                      InputLimitSwitchClosed := "20_TANKS_IP_DATA".RIO_05.SECOND_TANK.TANK_VENT_A_CLSD,
                      Open => "1092_HMI_OP_FLAGS".CV427_428_PVVA_Alarms[11].Open,
                      Closed => "1092_HMI_OP_FLAGS".CV427_428_PVVA_Alarms[11].Closed,
                      Moving => "1092_HMI_OP_FLAGS".CV427_428_PVVA_Alarms[11].Moving,
                      Fault => "1092_HMI_OP_FLAGS".CV427_428_PVVA_Alarms[11].Fault);
END_REGION

REGION Network 6: 600-CV-427, 600-CV-428 Alarms (RIO 06: 6P, 6S)
   RUNG wire#powerrail
      "1603_VALVE_STATE"(InputLimitSwitchOpen := "20_TANKS_IP_DATA".RIO_06.FIRST_TANK.TANK_VENT_A_OPEN, InputLimitSwitchClosed := "20_TANKS_IP_DATA".RIO_06.FIRST_TANK.TANK_VENT_A_CLSD, Open => "1092_HMI_OP_FLAGS".CV427_428_PVVA_Alarms[12].Open, Closed => "1092_HMI_OP_FLAGS".CV427_428_PVVA_Alarms[12].Closed, Moving => "1092_HMI_OP_FLAGS".CV427_428_PVVA_Alarms[12].Moving, Fault => "1092_HMI_OP_FLAGS".CV427_428_PVVA_Alarms[12].Fault)
   END_RUNG
   RUNG wire#powerrail
      "1603_VALVE_STATE"(InputLimitSwitchOpen := "20_TANKS_IP_DATA".RIO_06.SECOND_TANK.TANK_VENT_A_OPEN, InputLimitSwitchClosed := "20_TANKS_IP_DATA".RIO_06.SECOND_TANK.TANK_VENT_A_CLSD, Open => "1092_HMI_OP_FLAGS".CV427_428_PVVA_Alarms[13].Open, Closed => "1092_HMI_OP_FLAGS".CV427_428_PVVA_Alarms[13].Closed, Moving => "1092_HMI_OP_FLAGS".CV427_428_PVVA_Alarms[13].Moving, Fault => "1092_HMI_OP_FLAGS".CV427_428_PVVA_Alarms[13].Fault)
   END_RUNG
   // the same network as SCL:
   "1603_VALVE_STATE"(InputLimitSwitchOpen := "20_TANKS_IP_DATA".RIO_06.FIRST_TANK.TANK_VENT_A_OPEN,
                      InputLimitSwitchClosed := "20_TANKS_IP_DATA".RIO_06.FIRST_TANK.TANK_VENT_A_CLSD,
                      Open => "1092_HMI_OP_FLAGS".CV427_428_PVVA_Alarms[12].Open,
                      Closed => "1092_HMI_OP_FLAGS".CV427_428_PVVA_Alarms[12].Closed,
                      Moving => "1092_HMI_OP_FLAGS".CV427_428_PVVA_Alarms[12].Moving,
                      Fault => "1092_HMI_OP_FLAGS".CV427_428_PVVA_Alarms[12].Fault);
   "1603_VALVE_STATE"(InputLimitSwitchOpen := "20_TANKS_IP_DATA".RIO_06.SECOND_TANK.TANK_VENT_A_OPEN,
                      InputLimitSwitchClosed := "20_TANKS_IP_DATA".RIO_06.SECOND_TANK.TANK_VENT_A_CLSD,
                      Open => "1092_HMI_OP_FLAGS".CV427_428_PVVA_Alarms[13].Open,
                      Closed => "1092_HMI_OP_FLAGS".CV427_428_PVVA_Alarms[13].Closed,
                      Moving => "1092_HMI_OP_FLAGS".CV427_428_PVVA_Alarms[13].Moving,
                      Fault => "1092_HMI_OP_FLAGS".CV427_428_PVVA_Alarms[13].Fault);
END_REGION

REGION Network 7: 600-CV-427, 600-CV-428 Alarms (RIO 07: APT)
   RUNG wire#powerrail
      "1603_VALVE_STATE"(InputLimitSwitchOpen := "20_TANKS_IP_DATA".RIO_07.FIRST_TANK.TANK_VENT_A_OPEN, InputLimitSwitchClosed := "20_TANKS_IP_DATA".RIO_07.FIRST_TANK.TANK_VENT_A_CLSD, Open => "1092_HMI_OP_FLAGS".CV427_428_PVVA_Alarms[14].Open, Closed => "1092_HMI_OP_FLAGS".CV427_428_PVVA_Alarms[14].Closed, Moving => "1092_HMI_OP_FLAGS".CV427_428_PVVA_Alarms[14].Moving, Fault => "1092_HMI_OP_FLAGS".CV427_428_PVVA_Alarms[14].Fault)
   END_RUNG
   // the same network as SCL:
   "1603_VALVE_STATE"(InputLimitSwitchOpen := "20_TANKS_IP_DATA".RIO_07.FIRST_TANK.TANK_VENT_A_OPEN,
                      InputLimitSwitchClosed := "20_TANKS_IP_DATA".RIO_07.FIRST_TANK.TANK_VENT_A_CLSD,
                      Open => "1092_HMI_OP_FLAGS".CV427_428_PVVA_Alarms[14].Open,
                      Closed => "1092_HMI_OP_FLAGS".CV427_428_PVVA_Alarms[14].Closed,
                      Moving => "1092_HMI_OP_FLAGS".CV427_428_PVVA_Alarms[14].Moving,
                      Fault => "1092_HMI_OP_FLAGS".CV427_428_PVVA_Alarms[14].Fault);
END_REGION
END_FUNCTION

FUNCTION "1087_600CV429_430_STATUS" : Void   // FC1087, LAD
{ S7_Optimized_Access := 'TRUE' }
VERSION : 0.1
// Calculate the valve status' for each of the Vent B Valves.
BEGIN

REGION Network 1: 600-CV-429, 600-CV-430 Alarms (RIO 01: FPT. 1P, 1S)
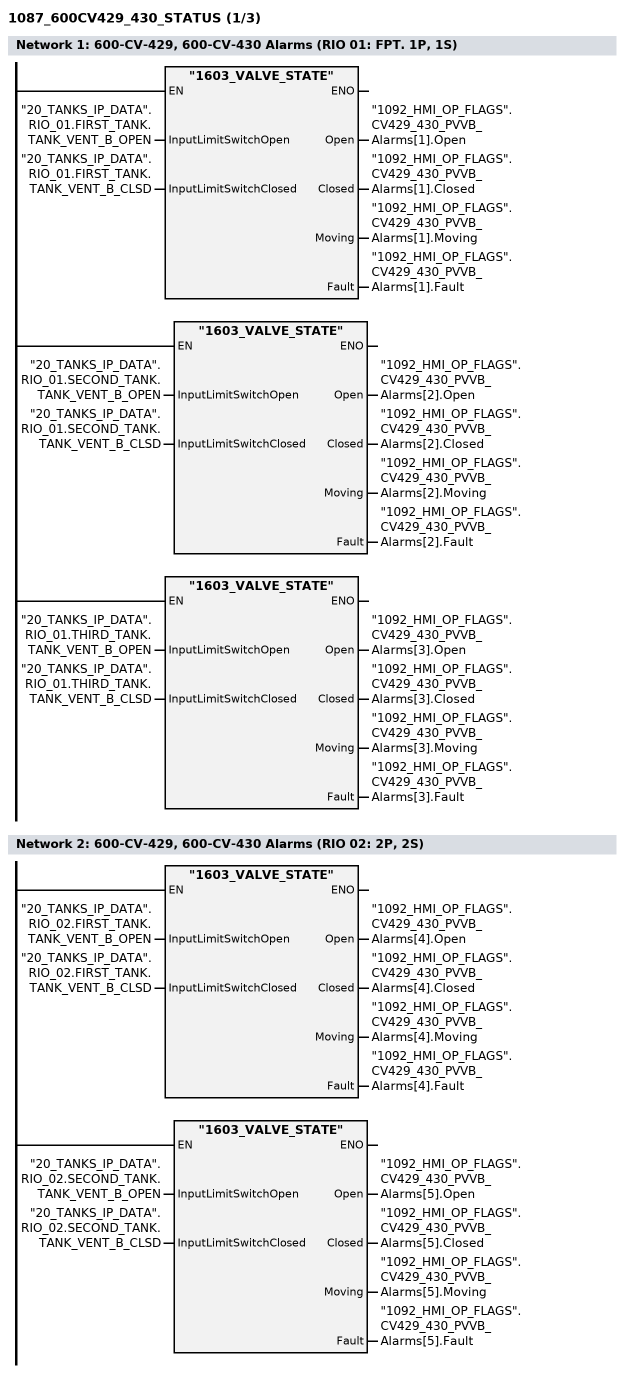
   RUNG wire#powerrail
      "1603_VALVE_STATE"(InputLimitSwitchOpen := "20_TANKS_IP_DATA".RIO_01.FIRST_TANK.TANK_VENT_B_OPEN, InputLimitSwitchClosed := "20_TANKS_IP_DATA".RIO_01.FIRST_TANK.TANK_VENT_B_CLSD, Open => "1092_HMI_OP_FLAGS".CV429_430_PVVB_Alarms[1].Open, Closed => "1092_HMI_OP_FLAGS".CV429_430_PVVB_Alarms[1].Closed, Moving => "1092_HMI_OP_FLAGS".CV429_430_PVVB_Alarms[1].Moving, Fault => "1092_HMI_OP_FLAGS".CV429_430_PVVB_Alarms[1].Fault)
   END_RUNG
   RUNG wire#powerrail
      "1603_VALVE_STATE"(InputLimitSwitchOpen := "20_TANKS_IP_DATA".RIO_01.SECOND_TANK.TANK_VENT_B_OPEN, InputLimitSwitchClosed := "20_TANKS_IP_DATA".RIO_01.SECOND_TANK.TANK_VENT_B_CLSD, Open => "1092_HMI_OP_FLAGS".CV429_430_PVVB_Alarms[2].Open, Closed => "1092_HMI_OP_FLAGS".CV429_430_PVVB_Alarms[2].Closed, Moving => "1092_HMI_OP_FLAGS".CV429_430_PVVB_Alarms[2].Moving, Fault => "1092_HMI_OP_FLAGS".CV429_430_PVVB_Alarms[2].Fault)
   END_RUNG
   RUNG wire#powerrail
      "1603_VALVE_STATE"(InputLimitSwitchOpen := "20_TANKS_IP_DATA".RIO_01.THIRD_TANK.TANK_VENT_B_OPEN, InputLimitSwitchClosed := "20_TANKS_IP_DATA".RIO_01.THIRD_TANK.TANK_VENT_B_CLSD, Open => "1092_HMI_OP_FLAGS".CV429_430_PVVB_Alarms[3].Open, Closed => "1092_HMI_OP_FLAGS".CV429_430_PVVB_Alarms[3].Closed, Moving => "1092_HMI_OP_FLAGS".CV429_430_PVVB_Alarms[3].Moving, Fault => "1092_HMI_OP_FLAGS".CV429_430_PVVB_Alarms[3].Fault)
   END_RUNG
   // the same network as SCL:
   "1603_VALVE_STATE"(InputLimitSwitchOpen := "20_TANKS_IP_DATA".RIO_01.FIRST_TANK.TANK_VENT_B_OPEN,
                      InputLimitSwitchClosed := "20_TANKS_IP_DATA".RIO_01.FIRST_TANK.TANK_VENT_B_CLSD,
                      Open => "1092_HMI_OP_FLAGS".CV429_430_PVVB_Alarms[1].Open,
                      Closed => "1092_HMI_OP_FLAGS".CV429_430_PVVB_Alarms[1].Closed,
                      Moving => "1092_HMI_OP_FLAGS".CV429_430_PVVB_Alarms[1].Moving,
                      Fault => "1092_HMI_OP_FLAGS".CV429_430_PVVB_Alarms[1].Fault);
   "1603_VALVE_STATE"(InputLimitSwitchOpen := "20_TANKS_IP_DATA".RIO_01.SECOND_TANK.TANK_VENT_B_OPEN,
                      InputLimitSwitchClosed := "20_TANKS_IP_DATA".RIO_01.SECOND_TANK.TANK_VENT_B_CLSD,
                      Open => "1092_HMI_OP_FLAGS".CV429_430_PVVB_Alarms[2].Open,
                      Closed => "1092_HMI_OP_FLAGS".CV429_430_PVVB_Alarms[2].Closed,
                      Moving => "1092_HMI_OP_FLAGS".CV429_430_PVVB_Alarms[2].Moving,
                      Fault => "1092_HMI_OP_FLAGS".CV429_430_PVVB_Alarms[2].Fault);
   "1603_VALVE_STATE"(InputLimitSwitchOpen := "20_TANKS_IP_DATA".RIO_01.THIRD_TANK.TANK_VENT_B_OPEN,
                      InputLimitSwitchClosed := "20_TANKS_IP_DATA".RIO_01.THIRD_TANK.TANK_VENT_B_CLSD,
                      Open => "1092_HMI_OP_FLAGS".CV429_430_PVVB_Alarms[3].Open,
                      Closed => "1092_HMI_OP_FLAGS".CV429_430_PVVB_Alarms[3].Closed,
                      Moving => "1092_HMI_OP_FLAGS".CV429_430_PVVB_Alarms[3].Moving,
                      Fault => "1092_HMI_OP_FLAGS".CV429_430_PVVB_Alarms[3].Fault);
END_REGION

REGION Network 2: 600-CV-429, 600-CV-430 Alarms (RIO 02: 2P, 2S)
   RUNG wire#powerrail
      "1603_VALVE_STATE"(InputLimitSwitchOpen := "20_TANKS_IP_DATA".RIO_02.FIRST_TANK.TANK_VENT_B_OPEN, InputLimitSwitchClosed := "20_TANKS_IP_DATA".RIO_02.FIRST_TANK.TANK_VENT_B_CLSD, Open => "1092_HMI_OP_FLAGS".CV429_430_PVVB_Alarms[4].Open, Closed => "1092_HMI_OP_FLAGS".CV429_430_PVVB_Alarms[4].Closed, Moving => "1092_HMI_OP_FLAGS".CV429_430_PVVB_Alarms[4].Moving, Fault => "1092_HMI_OP_FLAGS".CV429_430_PVVB_Alarms[4].Fault)
   END_RUNG
   RUNG wire#powerrail
      "1603_VALVE_STATE"(InputLimitSwitchOpen := "20_TANKS_IP_DATA".RIO_02.SECOND_TANK.TANK_VENT_B_OPEN, InputLimitSwitchClosed := "20_TANKS_IP_DATA".RIO_02.SECOND_TANK.TANK_VENT_B_CLSD, Open => "1092_HMI_OP_FLAGS".CV429_430_PVVB_Alarms[5].Open, Closed => "1092_HMI_OP_FLAGS".CV429_430_PVVB_Alarms[5].Closed, Moving => "1092_HMI_OP_FLAGS".CV429_430_PVVB_Alarms[5].Moving, Fault => "1092_HMI_OP_FLAGS".CV429_430_PVVB_Alarms[5].Fault)
   END_RUNG
   // the same network as SCL:
   "1603_VALVE_STATE"(InputLimitSwitchOpen := "20_TANKS_IP_DATA".RIO_02.FIRST_TANK.TANK_VENT_B_OPEN,
                      InputLimitSwitchClosed := "20_TANKS_IP_DATA".RIO_02.FIRST_TANK.TANK_VENT_B_CLSD,
                      Open => "1092_HMI_OP_FLAGS".CV429_430_PVVB_Alarms[4].Open,
                      Closed => "1092_HMI_OP_FLAGS".CV429_430_PVVB_Alarms[4].Closed,
                      Moving => "1092_HMI_OP_FLAGS".CV429_430_PVVB_Alarms[4].Moving,
                      Fault => "1092_HMI_OP_FLAGS".CV429_430_PVVB_Alarms[4].Fault);
   "1603_VALVE_STATE"(InputLimitSwitchOpen := "20_TANKS_IP_DATA".RIO_02.SECOND_TANK.TANK_VENT_B_OPEN,
                      InputLimitSwitchClosed := "20_TANKS_IP_DATA".RIO_02.SECOND_TANK.TANK_VENT_B_CLSD,
                      Open => "1092_HMI_OP_FLAGS".CV429_430_PVVB_Alarms[5].Open,
                      Closed => "1092_HMI_OP_FLAGS".CV429_430_PVVB_Alarms[5].Closed,
                      Moving => "1092_HMI_OP_FLAGS".CV429_430_PVVB_Alarms[5].Moving,
                      Fault => "1092_HMI_OP_FLAGS".CV429_430_PVVB_Alarms[5].Fault);
END_REGION

REGION Network 3: 600-CV-429, 600-CV-430 Alarms (RIO 03: 3P, 3S)
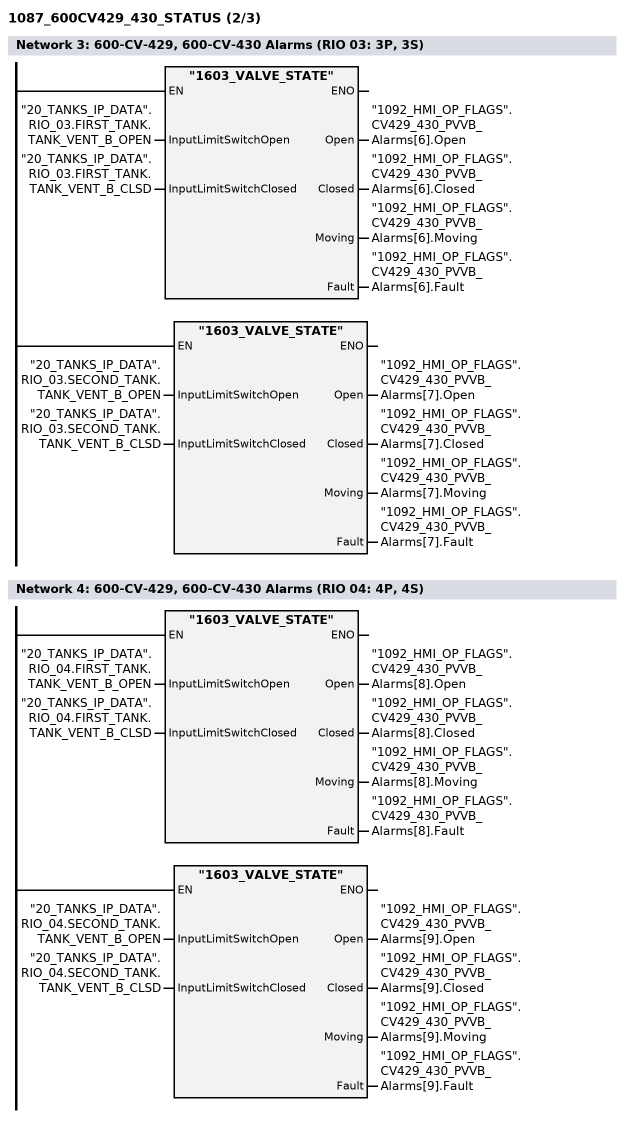
   RUNG wire#powerrail
      "1603_VALVE_STATE"(InputLimitSwitchOpen := "20_TANKS_IP_DATA".RIO_03.FIRST_TANK.TANK_VENT_B_OPEN, InputLimitSwitchClosed := "20_TANKS_IP_DATA".RIO_03.FIRST_TANK.TANK_VENT_B_CLSD, Open => "1092_HMI_OP_FLAGS".CV429_430_PVVB_Alarms[6].Open, Closed => "1092_HMI_OP_FLAGS".CV429_430_PVVB_Alarms[6].Closed, Moving => "1092_HMI_OP_FLAGS".CV429_430_PVVB_Alarms[6].Moving, Fault => "1092_HMI_OP_FLAGS".CV429_430_PVVB_Alarms[6].Fault)
   END_RUNG
   RUNG wire#powerrail
      "1603_VALVE_STATE"(InputLimitSwitchOpen := "20_TANKS_IP_DATA".RIO_03.SECOND_TANK.TANK_VENT_B_OPEN, InputLimitSwitchClosed := "20_TANKS_IP_DATA".RIO_03.SECOND_TANK.TANK_VENT_B_CLSD, Open => "1092_HMI_OP_FLAGS".CV429_430_PVVB_Alarms[7].Open, Closed => "1092_HMI_OP_FLAGS".CV429_430_PVVB_Alarms[7].Closed, Moving => "1092_HMI_OP_FLAGS".CV429_430_PVVB_Alarms[7].Moving, Fault => "1092_HMI_OP_FLAGS".CV429_430_PVVB_Alarms[7].Fault)
   END_RUNG
   // the same network as SCL:
   "1603_VALVE_STATE"(InputLimitSwitchOpen := "20_TANKS_IP_DATA".RIO_03.FIRST_TANK.TANK_VENT_B_OPEN,
                      InputLimitSwitchClosed := "20_TANKS_IP_DATA".RIO_03.FIRST_TANK.TANK_VENT_B_CLSD,
                      Open => "1092_HMI_OP_FLAGS".CV429_430_PVVB_Alarms[6].Open,
                      Closed => "1092_HMI_OP_FLAGS".CV429_430_PVVB_Alarms[6].Closed,
                      Moving => "1092_HMI_OP_FLAGS".CV429_430_PVVB_Alarms[6].Moving,
                      Fault => "1092_HMI_OP_FLAGS".CV429_430_PVVB_Alarms[6].Fault);
   "1603_VALVE_STATE"(InputLimitSwitchOpen := "20_TANKS_IP_DATA".RIO_03.SECOND_TANK.TANK_VENT_B_OPEN,
                      InputLimitSwitchClosed := "20_TANKS_IP_DATA".RIO_03.SECOND_TANK.TANK_VENT_B_CLSD,
                      Open => "1092_HMI_OP_FLAGS".CV429_430_PVVB_Alarms[7].Open,
                      Closed => "1092_HMI_OP_FLAGS".CV429_430_PVVB_Alarms[7].Closed,
                      Moving => "1092_HMI_OP_FLAGS".CV429_430_PVVB_Alarms[7].Moving,
                      Fault => "1092_HMI_OP_FLAGS".CV429_430_PVVB_Alarms[7].Fault);
END_REGION

REGION Network 4: 600-CV-429, 600-CV-430 Alarms (RIO 04: 4P, 4S)
   RUNG wire#powerrail
      "1603_VALVE_STATE"(InputLimitSwitchOpen := "20_TANKS_IP_DATA".RIO_04.FIRST_TANK.TANK_VENT_B_OPEN, InputLimitSwitchClosed := "20_TANKS_IP_DATA".RIO_04.FIRST_TANK.TANK_VENT_B_CLSD, Open => "1092_HMI_OP_FLAGS".CV429_430_PVVB_Alarms[8].Open, Closed => "1092_HMI_OP_FLAGS".CV429_430_PVVB_Alarms[8].Closed, Moving => "1092_HMI_OP_FLAGS".CV429_430_PVVB_Alarms[8].Moving, Fault => "1092_HMI_OP_FLAGS".CV429_430_PVVB_Alarms[8].Fault)
   END_RUNG
   RUNG wire#powerrail
      "1603_VALVE_STATE"(InputLimitSwitchOpen := "20_TANKS_IP_DATA".RIO_04.SECOND_TANK.TANK_VENT_B_OPEN, InputLimitSwitchClosed := "20_TANKS_IP_DATA".RIO_04.SECOND_TANK.TANK_VENT_B_CLSD, Open => "1092_HMI_OP_FLAGS".CV429_430_PVVB_Alarms[9].Open, Closed => "1092_HMI_OP_FLAGS".CV429_430_PVVB_Alarms[9].Closed, Moving => "1092_HMI_OP_FLAGS".CV429_430_PVVB_Alarms[9].Moving, Fault => "1092_HMI_OP_FLAGS".CV429_430_PVVB_Alarms[9].Fault)
   END_RUNG
   // the same network as SCL:
   "1603_VALVE_STATE"(InputLimitSwitchOpen := "20_TANKS_IP_DATA".RIO_04.FIRST_TANK.TANK_VENT_B_OPEN,
                      InputLimitSwitchClosed := "20_TANKS_IP_DATA".RIO_04.FIRST_TANK.TANK_VENT_B_CLSD,
                      Open => "1092_HMI_OP_FLAGS".CV429_430_PVVB_Alarms[8].Open,
                      Closed => "1092_HMI_OP_FLAGS".CV429_430_PVVB_Alarms[8].Closed,
                      Moving => "1092_HMI_OP_FLAGS".CV429_430_PVVB_Alarms[8].Moving,
                      Fault => "1092_HMI_OP_FLAGS".CV429_430_PVVB_Alarms[8].Fault);
   "1603_VALVE_STATE"(InputLimitSwitchOpen := "20_TANKS_IP_DATA".RIO_04.SECOND_TANK.TANK_VENT_B_OPEN,
                      InputLimitSwitchClosed := "20_TANKS_IP_DATA".RIO_04.SECOND_TANK.TANK_VENT_B_CLSD,
                      Open => "1092_HMI_OP_FLAGS".CV429_430_PVVB_Alarms[9].Open,
                      Closed => "1092_HMI_OP_FLAGS".CV429_430_PVVB_Alarms[9].Closed,
                      Moving => "1092_HMI_OP_FLAGS".CV429_430_PVVB_Alarms[9].Moving,
                      Fault => "1092_HMI_OP_FLAGS".CV429_430_PVVB_Alarms[9].Fault);
END_REGION

REGION Network 5: 600-CV-429, 600-CV-430 Alarms (RIO 05: 5P, 5S)
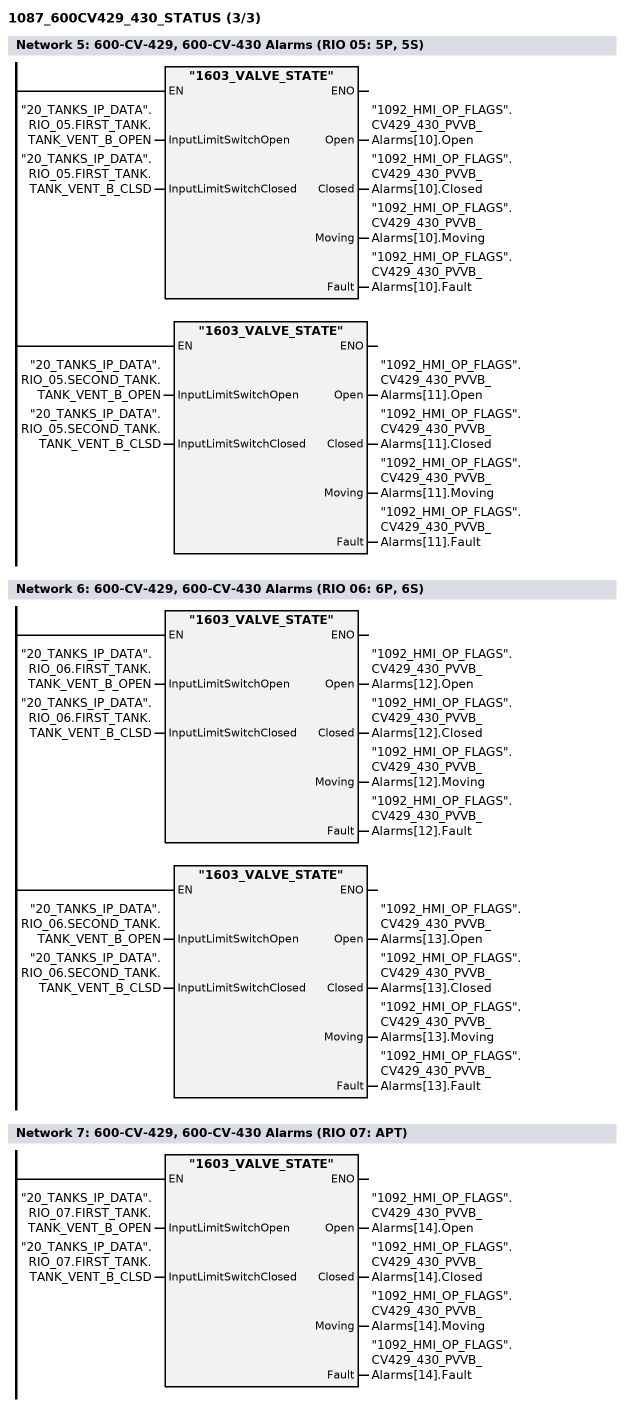
   RUNG wire#powerrail
      "1603_VALVE_STATE"(InputLimitSwitchOpen := "20_TANKS_IP_DATA".RIO_05.FIRST_TANK.TANK_VENT_B_OPEN, InputLimitSwitchClosed := "20_TANKS_IP_DATA".RIO_05.FIRST_TANK.TANK_VENT_B_CLSD, Open => "1092_HMI_OP_FLAGS".CV429_430_PVVB_Alarms[10].Open, Closed => "1092_HMI_OP_FLAGS".CV429_430_PVVB_Alarms[10].Closed, Moving => "1092_HMI_OP_FLAGS".CV429_430_PVVB_Alarms[10].Moving, Fault => "1092_HMI_OP_FLAGS".CV429_430_PVVB_Alarms[10].Fault)
   END_RUNG
   RUNG wire#powerrail
      "1603_VALVE_STATE"(InputLimitSwitchOpen := "20_TANKS_IP_DATA".RIO_05.SECOND_TANK.TANK_VENT_B_OPEN, InputLimitSwitchClosed := "20_TANKS_IP_DATA".RIO_05.SECOND_TANK.TANK_VENT_B_CLSD, Open => "1092_HMI_OP_FLAGS".CV429_430_PVVB_Alarms[11].Open, Closed => "1092_HMI_OP_FLAGS".CV429_430_PVVB_Alarms[11].Closed, Moving => "1092_HMI_OP_FLAGS".CV429_430_PVVB_Alarms[11].Moving, Fault => "1092_HMI_OP_FLAGS".CV429_430_PVVB_Alarms[11].Fault)
   END_RUNG
   // the same network as SCL:
   "1603_VALVE_STATE"(InputLimitSwitchOpen := "20_TANKS_IP_DATA".RIO_05.FIRST_TANK.TANK_VENT_B_OPEN,
                      InputLimitSwitchClosed := "20_TANKS_IP_DATA".RIO_05.FIRST_TANK.TANK_VENT_B_CLSD,
                      Open => "1092_HMI_OP_FLAGS".CV429_430_PVVB_Alarms[10].Open,
                      Closed => "1092_HMI_OP_FLAGS".CV429_430_PVVB_Alarms[10].Closed,
                      Moving => "1092_HMI_OP_FLAGS".CV429_430_PVVB_Alarms[10].Moving,
                      Fault => "1092_HMI_OP_FLAGS".CV429_430_PVVB_Alarms[10].Fault);
   "1603_VALVE_STATE"(InputLimitSwitchOpen := "20_TANKS_IP_DATA".RIO_05.SECOND_TANK.TANK_VENT_B_OPEN,
                      InputLimitSwitchClosed := "20_TANKS_IP_DATA".RIO_05.SECOND_TANK.TANK_VENT_B_CLSD,
                      Open => "1092_HMI_OP_FLAGS".CV429_430_PVVB_Alarms[11].Open,
                      Closed => "1092_HMI_OP_FLAGS".CV429_430_PVVB_Alarms[11].Closed,
                      Moving => "1092_HMI_OP_FLAGS".CV429_430_PVVB_Alarms[11].Moving,
                      Fault => "1092_HMI_OP_FLAGS".CV429_430_PVVB_Alarms[11].Fault);
END_REGION

REGION Network 6: 600-CV-429, 600-CV-430 Alarms (RIO 06: 6P, 6S)
   RUNG wire#powerrail
      "1603_VALVE_STATE"(InputLimitSwitchOpen := "20_TANKS_IP_DATA".RIO_06.FIRST_TANK.TANK_VENT_B_OPEN, InputLimitSwitchClosed := "20_TANKS_IP_DATA".RIO_06.FIRST_TANK.TANK_VENT_B_CLSD, Open => "1092_HMI_OP_FLAGS".CV429_430_PVVB_Alarms[12].Open, Closed => "1092_HMI_OP_FLAGS".CV429_430_PVVB_Alarms[12].Closed, Moving => "1092_HMI_OP_FLAGS".CV429_430_PVVB_Alarms[12].Moving, Fault => "1092_HMI_OP_FLAGS".CV429_430_PVVB_Alarms[12].Fault)
   END_RUNG
   RUNG wire#powerrail
      "1603_VALVE_STATE"(InputLimitSwitchOpen := "20_TANKS_IP_DATA".RIO_06.SECOND_TANK.TANK_VENT_B_OPEN, InputLimitSwitchClosed := "20_TANKS_IP_DATA".RIO_06.SECOND_TANK.TANK_VENT_B_CLSD, Open => "1092_HMI_OP_FLAGS".CV429_430_PVVB_Alarms[13].Open, Closed => "1092_HMI_OP_FLAGS".CV429_430_PVVB_Alarms[13].Closed, Moving => "1092_HMI_OP_FLAGS".CV429_430_PVVB_Alarms[13].Moving, Fault => "1092_HMI_OP_FLAGS".CV429_430_PVVB_Alarms[13].Fault)
   END_RUNG
   // the same network as SCL:
   "1603_VALVE_STATE"(InputLimitSwitchOpen := "20_TANKS_IP_DATA".RIO_06.FIRST_TANK.TANK_VENT_B_OPEN,
                      InputLimitSwitchClosed := "20_TANKS_IP_DATA".RIO_06.FIRST_TANK.TANK_VENT_B_CLSD,
                      Open => "1092_HMI_OP_FLAGS".CV429_430_PVVB_Alarms[12].Open,
                      Closed => "1092_HMI_OP_FLAGS".CV429_430_PVVB_Alarms[12].Closed,
                      Moving => "1092_HMI_OP_FLAGS".CV429_430_PVVB_Alarms[12].Moving,
                      Fault => "1092_HMI_OP_FLAGS".CV429_430_PVVB_Alarms[12].Fault);
   "1603_VALVE_STATE"(InputLimitSwitchOpen := "20_TANKS_IP_DATA".RIO_06.SECOND_TANK.TANK_VENT_B_OPEN,
                      InputLimitSwitchClosed := "20_TANKS_IP_DATA".RIO_06.SECOND_TANK.TANK_VENT_B_CLSD,
                      Open => "1092_HMI_OP_FLAGS".CV429_430_PVVB_Alarms[13].Open,
                      Closed => "1092_HMI_OP_FLAGS".CV429_430_PVVB_Alarms[13].Closed,
                      Moving => "1092_HMI_OP_FLAGS".CV429_430_PVVB_Alarms[13].Moving,
                      Fault => "1092_HMI_OP_FLAGS".CV429_430_PVVB_Alarms[13].Fault);
END_REGION

REGION Network 7: 600-CV-429, 600-CV-430 Alarms (RIO 07: APT)
   RUNG wire#powerrail
      "1603_VALVE_STATE"(InputLimitSwitchOpen := "20_TANKS_IP_DATA".RIO_07.FIRST_TANK.TANK_VENT_B_OPEN, InputLimitSwitchClosed := "20_TANKS_IP_DATA".RIO_07.FIRST_TANK.TANK_VENT_B_CLSD, Open => "1092_HMI_OP_FLAGS".CV429_430_PVVB_Alarms[14].Open, Closed => "1092_HMI_OP_FLAGS".CV429_430_PVVB_Alarms[14].Closed, Moving => "1092_HMI_OP_FLAGS".CV429_430_PVVB_Alarms[14].Moving, Fault => "1092_HMI_OP_FLAGS".CV429_430_PVVB_Alarms[14].Fault)
   END_RUNG
   // the same network as SCL:
   "1603_VALVE_STATE"(InputLimitSwitchOpen := "20_TANKS_IP_DATA".RIO_07.FIRST_TANK.TANK_VENT_B_OPEN,
                      InputLimitSwitchClosed := "20_TANKS_IP_DATA".RIO_07.FIRST_TANK.TANK_VENT_B_CLSD,
                      Open => "1092_HMI_OP_FLAGS".CV429_430_PVVB_Alarms[14].Open,
                      Closed => "1092_HMI_OP_FLAGS".CV429_430_PVVB_Alarms[14].Closed,
                      Moving => "1092_HMI_OP_FLAGS".CV429_430_PVVB_Alarms[14].Moving,
                      Fault => "1092_HMI_OP_FLAGS".CV429_430_PVVB_Alarms[14].Fault);
END_REGION
END_FUNCTION

// folder: 1000 - 1999 BWT System Control/1100 - 1104 BWTS Control

